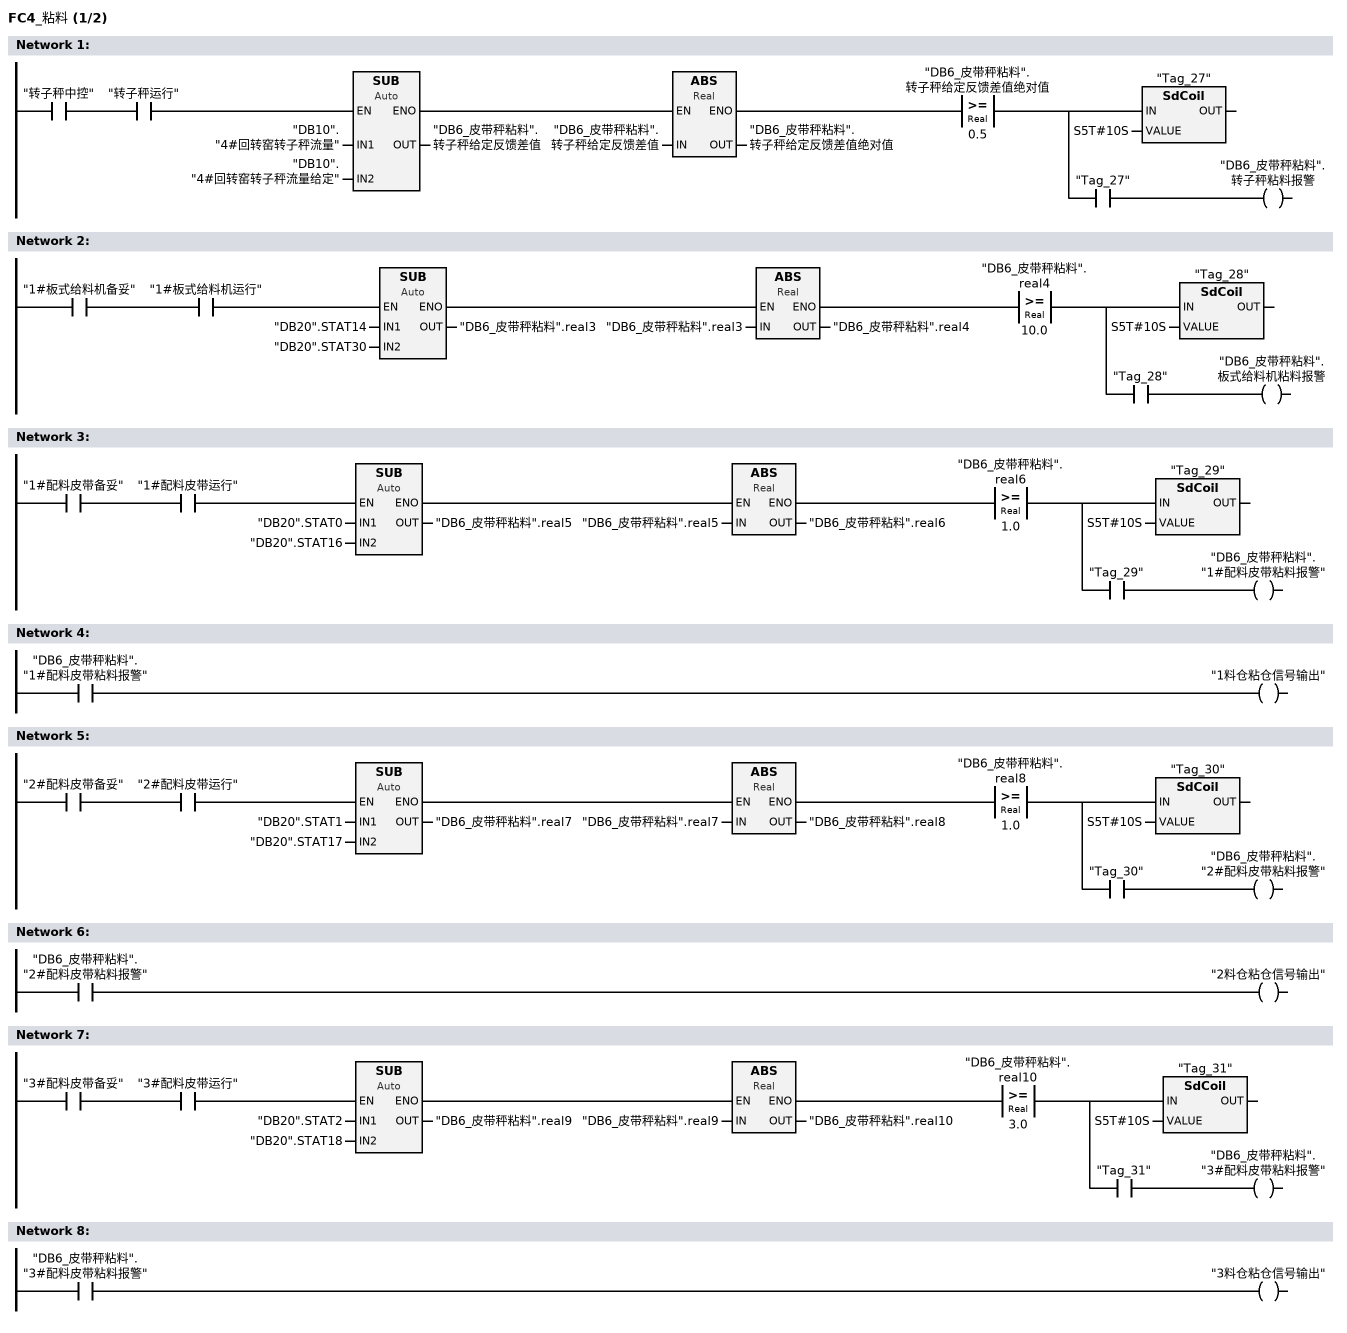
   // no SCL statement known for SdCoil: written as a call
   #_w1 := "转子秤中控" AND "转子秤运行";
   IF #_w1 THEN
       "DB6_皮带秤粘料".转子秤给定反馈差值 := "DB10"."4#回转窑转子秤流量" - "DB10"."4#回转窑转子秤流量给定";
       "DB6_皮带秤粘料".转子秤给定反馈差值绝对值 := ABS("DB6_皮带秤粘料".转子秤给定反馈差值);
   END_IF;
   #_w2 := #_w1 AND ("DB6_皮带秤粘料".转子秤给定反馈差值绝对值 >= 0.5);
   SdCoil(in := #_w2, value := S5T#10S, operand := "Tag_27");
   "DB6_皮带秤粘料".转子秤粘料报警 := #_w2 AND "Tag_27";
END_REGION

REGION Network 2
   // no SCL statement known for SdCoil: written as a call
   #_w1 := "1#板式给料机备妥" AND "1#板式给料机运行";
   IF #_w1 THEN
       "DB6_皮带秤粘料".real3 := "DB20".STAT14 - "DB20".STAT30;
       "DB6_皮带秤粘料".real4 := ABS("DB6_皮带秤粘料".real3);
   END_IF;
   #_w2 := #_w1 AND ("DB6_皮带秤粘料".real4 >= 10.0);
   SdCoil(in := #_w2, value := S5T#10S, operand := "Tag_28");
   "DB6_皮带秤粘料".板式给料机粘料报警 := #_w2 AND "Tag_28";
END_REGION

REGION Network 3
   // no SCL statement known for SdCoil: written as a call
   #_w1 := "1#配料皮带备妥" AND "1#配料皮带运行";
   IF #_w1 THEN
       "DB6_皮带秤粘料".real5 := "DB20".STAT0 - "DB20".STAT16;
       "DB6_皮带秤粘料".real6 := ABS("DB6_皮带秤粘料".real5);
   END_IF;
   #_w2 := #_w1 AND ("DB6_皮带秤粘料".real6 >= 1.0);
   SdCoil(in := #_w2, value := S5T#10S, operand := "Tag_29");
   "DB6_皮带秤粘料"."1#配料皮带粘料报警" := #_w2 AND "Tag_29";
END_REGION

REGION Network 4
   RUNG wire#powerrail
      Contact( "DB6_皮带秤粘料"."1#配料皮带粘料报警" )
      Coil( "1料仓粘仓信号输出" )
   END_RUNG
   // the same network as SCL:
   "1料仓粘仓信号输出" := "DB6_皮带秤粘料"."1#配料皮带粘料报警";
END_REGION

REGION Network 5
   // no SCL statement known for SdCoil: written as a call
   #_w1 := "2#配料皮带备妥" AND "2#配料皮带运行";
   IF #_w1 THEN
       "DB6_皮带秤粘料".real7 := "DB20".STAT1 - "DB20".STAT17;
       "DB6_皮带秤粘料".real8 := ABS("DB6_皮带秤粘料".real7);
   END_IF;
   #_w2 := #_w1 AND ("DB6_皮带秤粘料".real8 >= 1.0);
   SdCoil(in := #_w2, value := S5T#10S, operand := "Tag_30");
   "DB6_皮带秤粘料"."2#配料皮带粘料报警" := #_w2 AND "Tag_30";
END_REGION

REGION Network 6
   RUNG wire#powerrail
      Contact( "DB6_皮带秤粘料"."2#配料皮带粘料报警" )
      Coil( "2料仓粘仓信号输出" )
   END_RUNG
   // the same network as SCL:
   "2料仓粘仓信号输出" := "DB6_皮带秤粘料"."2#配料皮带粘料报警";
END_REGION

REGION Network 7
   // no SCL statement known for SdCoil: written as a call
   #_w1 := "3#配料皮带备妥" AND "3#配料皮带运行";
   IF #_w1 THEN
       "DB6_皮带秤粘料".real9 := "DB20".STAT2 - "DB20".STAT18;
       "DB6_皮带秤粘料".real10 := ABS("DB6_皮带秤粘料".real9);
   END_IF;
   #_w2 := #_w1 AND ("DB6_皮带秤粘料".real10 >= 3.0);
   SdCoil(in := #_w2, value := S5T#10S, operand := "Tag_31");
   "DB6_皮带秤粘料"."3#配料皮带粘料报警" := #_w2 AND "Tag_31";
END_REGION

REGION Network 8
   RUNG wire#powerrail
      Contact( "DB6_皮带秤粘料"."3#配料皮带粘料报警" )
      Coil( "3料仓粘仓信号输出" )
   END_RUNG
   // the same network as SCL:
   "3料仓粘仓信号输出" := "DB6_皮带秤粘料"."3#配料皮带粘料报警";
END_REGION

REGION Network 9
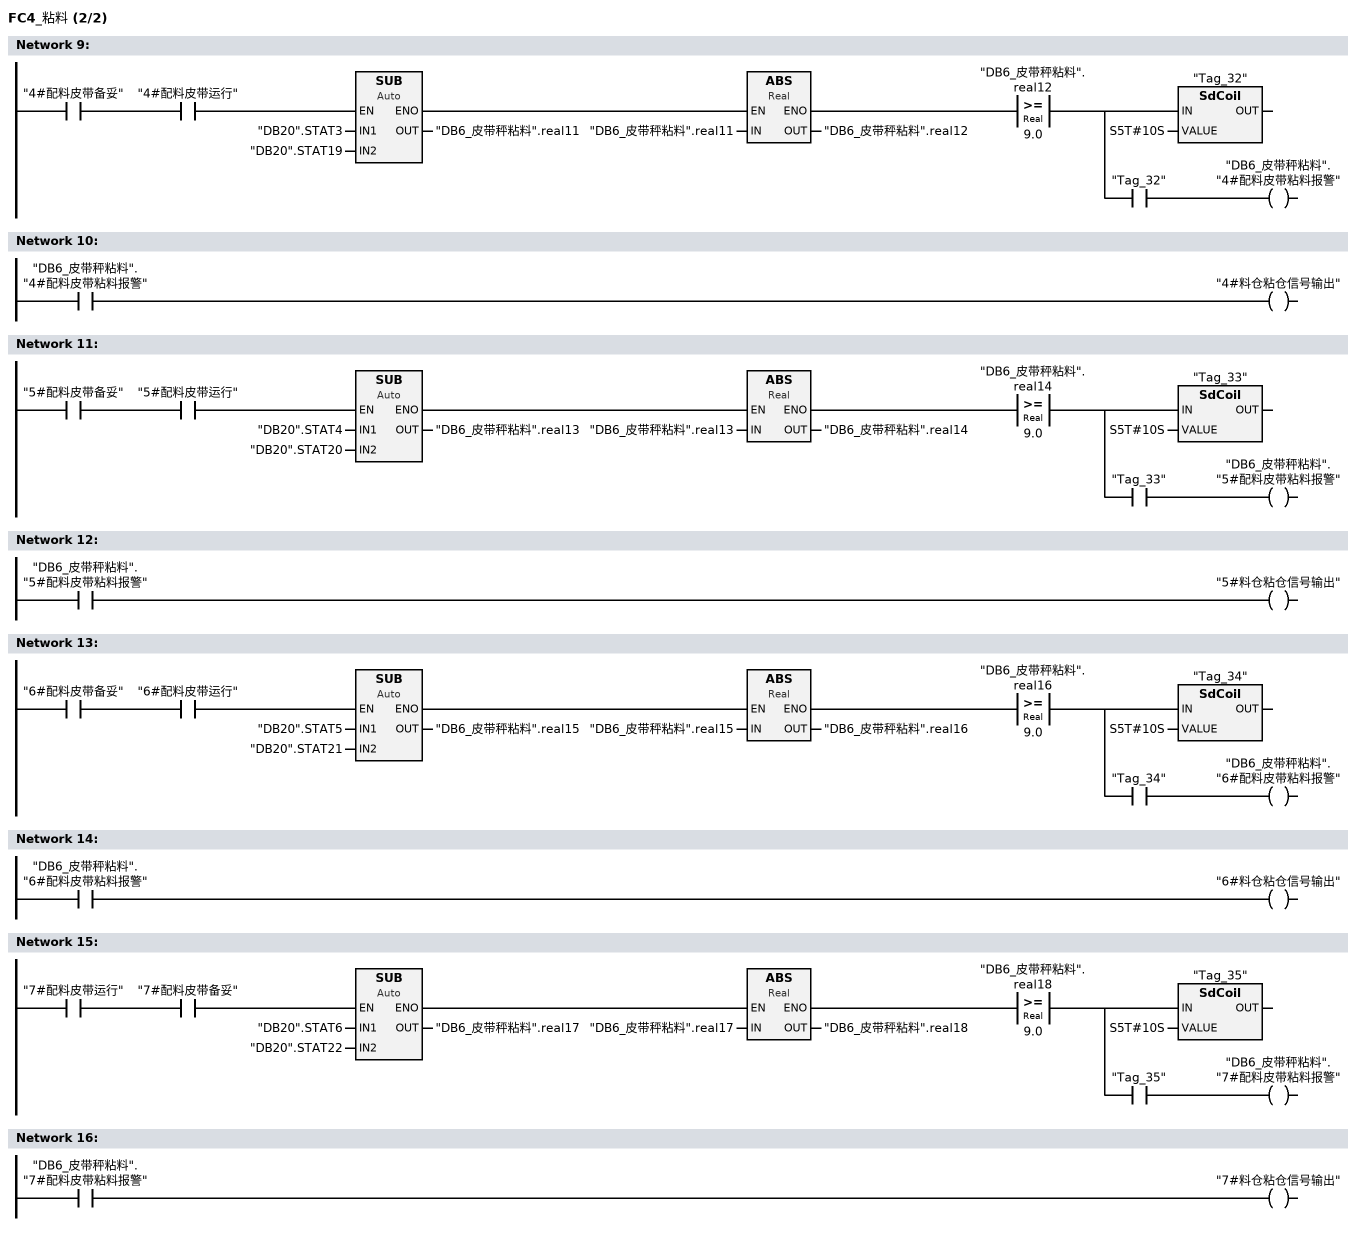
   // no SCL statement known for SdCoil: written as a call
   #_w1 := "4#配料皮带备妥" AND "4#配料皮带运行";
   IF #_w1 THEN
       "DB6_皮带秤粘料".real11 := "DB20".STAT3 - "DB20".STAT19;
       "DB6_皮带秤粘料".real12 := ABS("DB6_皮带秤粘料".real11);
   END_IF;
   #_w2 := #_w1 AND ("DB6_皮带秤粘料".real12 >= 9.0);
   SdCoil(in := #_w2, value := S5T#10S, operand := "Tag_32");
   "DB6_皮带秤粘料"."4#配料皮带粘料报警" := #_w2 AND "Tag_32";
END_REGION

REGION Network 10
   RUNG wire#powerrail
      Contact( "DB6_皮带秤粘料"."4#配料皮带粘料报警" )
      Coil( "4#料仓粘仓信号输出" )
   END_RUNG
   // the same network as SCL:
   "4#料仓粘仓信号输出" := "DB6_皮带秤粘料"."4#配料皮带粘料报警";
END_REGION

REGION Network 11
   // no SCL statement known for SdCoil: written as a call
   #_w1 := "5#配料皮带备妥" AND "5#配料皮带运行";
   IF #_w1 THEN
       "DB6_皮带秤粘料".real13 := "DB20".STAT4 - "DB20".STAT20;
       "DB6_皮带秤粘料".real14 := ABS("DB6_皮带秤粘料".real13);
   END_IF;
   #_w2 := #_w1 AND ("DB6_皮带秤粘料".real14 >= 9.0);
   SdCoil(in := #_w2, value := S5T#10S, operand := "Tag_33");
   "DB6_皮带秤粘料"."5#配料皮带粘料报警" := #_w2 AND "Tag_33";
END_REGION

REGION Network 12
   RUNG wire#powerrail
      Contact( "DB6_皮带秤粘料"."5#配料皮带粘料报警" )
      Coil( "5#料仓粘仓信号输出" )
   END_RUNG
   // the same network as SCL:
   "5#料仓粘仓信号输出" := "DB6_皮带秤粘料"."5#配料皮带粘料报警";
END_REGION

REGION Network 13
   // no SCL statement known for SdCoil: written as a call
   #_w1 := "6#配料皮带备妥" AND "6#配料皮带运行";
   IF #_w1 THEN
       "DB6_皮带秤粘料".real15 := "DB20".STAT5 - "DB20".STAT21;
       "DB6_皮带秤粘料".real16 := ABS("DB6_皮带秤粘料".real15);
   END_IF;
   #_w2 := #_w1 AND ("DB6_皮带秤粘料".real16 >= 9.0);
   SdCoil(in := #_w2, value := S5T#10S, operand := "Tag_34");
   "DB6_皮带秤粘料"."6#配料皮带粘料报警" := #_w2 AND "Tag_34";
END_REGION

REGION Network 14
   RUNG wire#powerrail
      Contact( "DB6_皮带秤粘料"."6#配料皮带粘料报警" )
      Coil( "6#料仓粘仓信号输出" )
   END_RUNG
   // the same network as SCL:
   "6#料仓粘仓信号输出" := "DB6_皮带秤粘料"."6#配料皮带粘料报警";
END_REGION

REGION Network 15
   // no SCL statement known for SdCoil: written as a call
   #_w1 := "7#配料皮带运行" AND "7#配料皮带备妥";
   IF #_w1 THEN
       "DB6_皮带秤粘料".real17 := "DB20".STAT6 - "DB20".STAT22;
       "DB6_皮带秤粘料".real18 := ABS("DB6_皮带秤粘料".real17);
   END_IF;
   #_w2 := #_w1 AND ("DB6_皮带秤粘料".real18 >= 9.0);
   SdCoil(in := #_w2, value := S5T#10S, operand := "Tag_35");
   "DB6_皮带秤粘料"."7#配料皮带粘料报警" := #_w2 AND "Tag_35";
END_REGION

REGION Network 16
   RUNG wire#powerrail
      Contact( "DB6_皮带秤粘料"."7#配料皮带粘料报警" )
      Coil( "7#料仓粘仓信号输出" )
   END_RUNG
   // the same network as SCL:
   "7#料仓粘仓信号输出" := "DB6_皮带秤粘料"."7#配料皮带粘料报警";
END_REGION
END_FUNCTION

FUNCTION "回转窑控制" : Void   // FC11, LAD
{ S7_Optimized_Access := 'FALSE' }
VERSION : 0.1
   VAR_TEMP   // added for the SCL form of the ladder/FBD networks
      _w1 : Bool;
      _s5time1 : S5Time;
   END_VAR
BEGIN

REGION Network 1
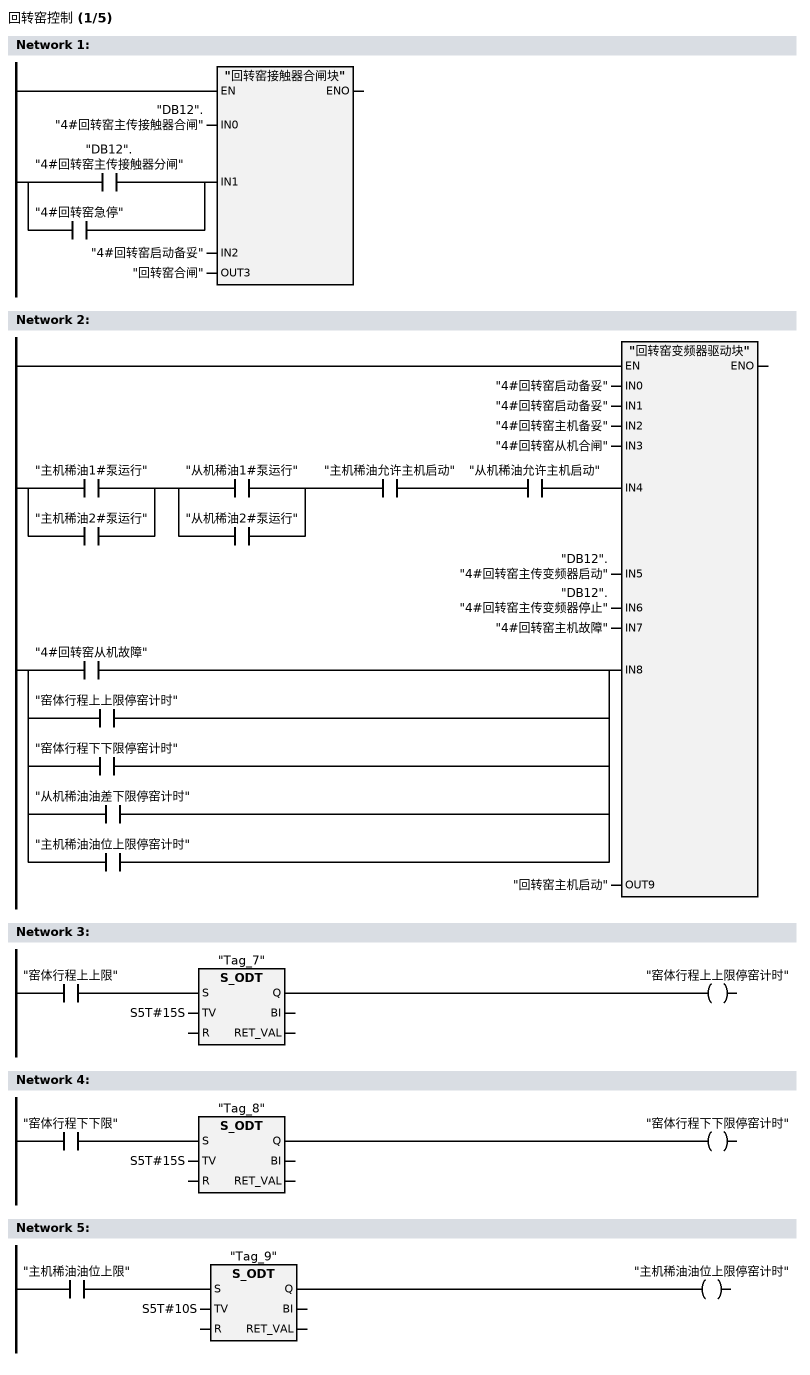
   RUNG wire#powerrail
      "回转窑接触器合闸块"(IN1 := wire#w1, IN0 := "DB12"."4#回转窑主传接触器合闸", IN2 := "4#回转窑启动备妥", OUT3 := "回转窑合闸")
   END_RUNG
   RUNG wire#powerrail
      Contact( "DB12"."4#回转窑主传接触器分闸" )
   END_RUNG wire#w1
   RUNG wire#powerrail
      Contact( "4#回转窑急停" )
   END_RUNG wire#w1
   // the same network as SCL:
   "回转窑接触器合闸块"(IN0 := "DB12"."4#回转窑主传接触器合闸",
               IN1 := "DB12"."4#回转窑主传接触器分闸" OR "4#回转窑急停",
               IN2 := "4#回转窑启动备妥",
               OUT3 := "回转窑合闸");
END_REGION

REGION Network 2
   RUNG wire#powerrail
      "回转窑变频器驱动块"(IN4 := wire#w3, IN8 := wire#w4, IN0 := "4#回转窑启动备妥", IN1 := "4#回转窑启动备妥", IN2 := "4#回转窑主机备妥", IN3 := "4#回转窑从机合闸", IN5 := "DB12"."4#回转窑主传变频器启动", IN6 := "DB12"."4#回转窑主传变频器停止", IN7 := "4#回转窑主机故障", OUT9 := "回转窑主机启动")
   END_RUNG
   RUNG wire#powerrail
      Contact( "主机稀油1#泵运行" )
      wire#w1
      Contact( "从机稀油1#泵运行" )
      wire#w2
      Contact( "主机稀油允许主机启动" )
      Contact( "从机稀油允许主机启动" )
   END_RUNG wire#w3
   RUNG wire#powerrail
      Contact( "主机稀油2#泵运行" )
   END_RUNG wire#w1
   RUNG wire#w1
      Contact( "从机稀油2#泵运行" )
   END_RUNG wire#w2
   RUNG wire#powerrail
      Contact( "4#回转窑从机故障" )
   END_RUNG wire#w4
   RUNG wire#powerrail
      Contact( "窑体行程上上限停窑计时" )
   END_RUNG wire#w4
   RUNG wire#powerrail
      Contact( "窑体行程下下限停窑计时" )
   END_RUNG wire#w4
   RUNG wire#powerrail
      Contact( "从机稀油油差下限停窑计时" )
   END_RUNG wire#w4
   RUNG wire#powerrail
      Contact( "主机稀油油位上限停窑计时" )
   END_RUNG wire#w4
   // the same network as SCL:
   "回转窑变频器驱动块"(IN0 := "4#回转窑启动备妥",
               IN1 := "4#回转窑启动备妥",
               IN2 := "4#回转窑主机备妥",
               IN3 := "4#回转窑从机合闸",
               IN4 := ("主机稀油1#泵运行" OR "主机稀油2#泵运行") AND ("从机稀油1#泵运行" OR "从机稀油2#泵运行") AND "主机稀油允许主机启动" AND "从机稀油允许主机启动",
               IN5 := "DB12"."4#回转窑主传变频器启动",
               IN6 := "DB12"."4#回转窑主传变频器停止",
               IN7 := "4#回转窑主机故障",
               IN8 := "4#回转窑从机故障" OR "窑体行程上上限停窑计时" OR "窑体行程下下限停窑计时" OR "从机稀油油差下限停窑计时" OR "主机稀油油位上限停窑计时",
               OUT9 := "回转窑主机启动");
END_REGION

REGION Network 3
   RUNG wire#powerrail
      Contact( "窑体行程上上限" )
      S_ODT(T_NO := "Tag_7", TV := S5T#15S, R :=, BI =>, RET_VAL =>)
      Coil( "窑体行程上上限停窑计时" )
   END_RUNG
   // the same network as SCL:
   #_s5time1 := S_ODT(T_NO := "Tag_7", TV := S5T#15S, S := "窑体行程上上限", Q => #_w1);
   "窑体行程上上限停窑计时" := #_w1;
END_REGION

REGION Network 4
   RUNG wire#powerrail
      Contact( "窑体行程下下限" )
      S_ODT(T_NO := "Tag_8", TV := S5T#15S, R :=, BI =>, RET_VAL =>)
      Coil( "窑体行程下下限停窑计时" )
   END_RUNG
   // the same network as SCL:
   #_s5time1 := S_ODT(T_NO := "Tag_8", TV := S5T#15S, S := "窑体行程下下限", Q => #_w1);
   "窑体行程下下限停窑计时" := #_w1;
END_REGION

REGION Network 5
   RUNG wire#powerrail
      Contact( "主机稀油油位上限" )
      S_ODT(T_NO := "Tag_9", TV := S5T#10S, R :=, BI =>, RET_VAL =>)
      Coil( "主机稀油油位上限停窑计时" )
   END_RUNG
   // the same network as SCL:
   #_s5time1 := S_ODT(T_NO := "Tag_9", S := "主机稀油油位上限", TV := S5T#10S, Q => #_w1);
   "主机稀油油位上限停窑计时" := #_w1;
END_REGION

REGION Network 6
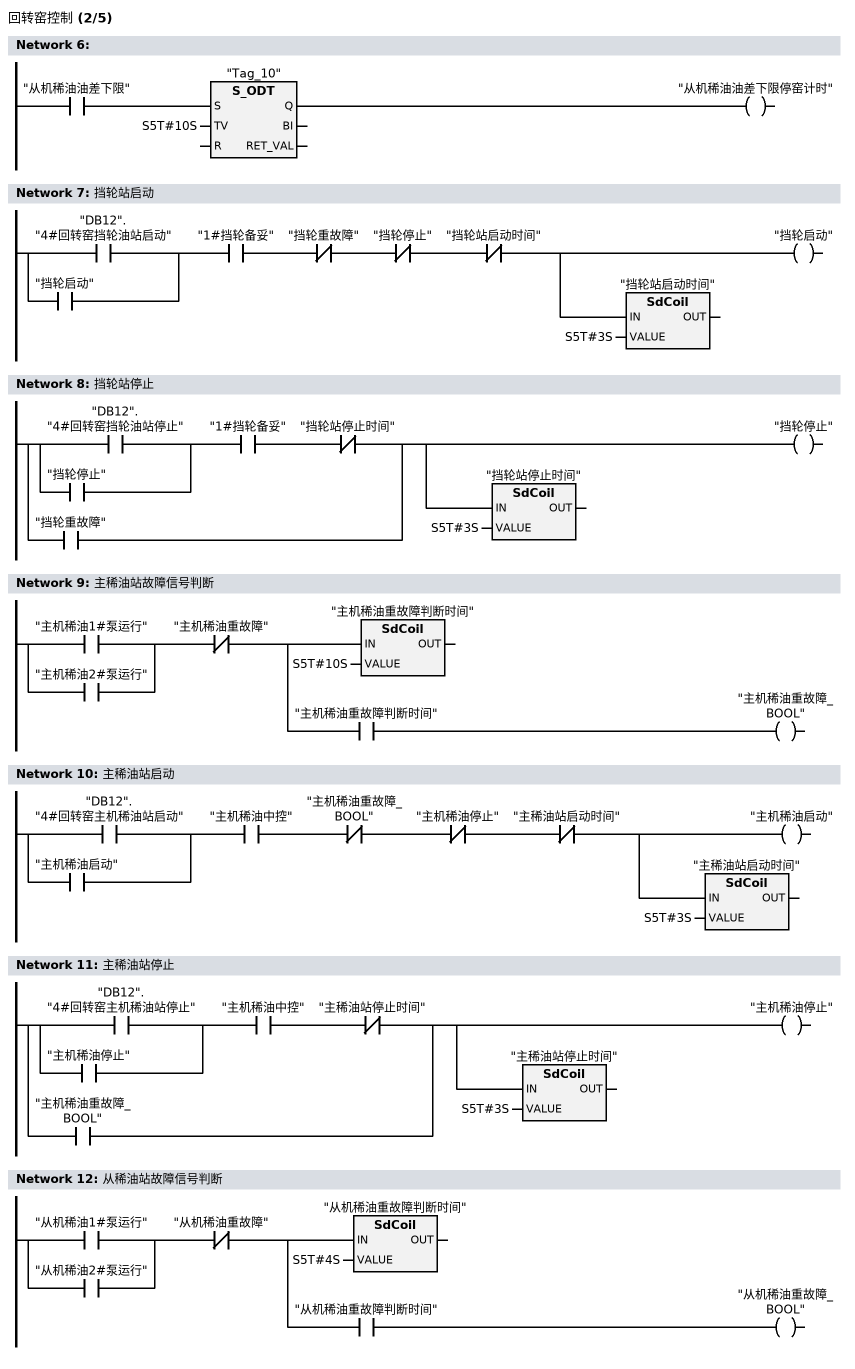
   RUNG wire#powerrail
      Contact( "从机稀油油差下限" )
      S_ODT(T_NO := "Tag_10", TV := S5T#10S, R :=, BI =>, RET_VAL =>)
      Coil( "从机稀油油差下限停窑计时" )
   END_RUNG
   // the same network as SCL:
   #_s5time1 := S_ODT(T_NO := "Tag_10", TV := S5T#10S, S := "从机稀油油差下限", Q => #_w1);
   "从机稀油油差下限停窑计时" := #_w1;
END_REGION

REGION Network 7: 挡轮站启动
   // no SCL statement known for SdCoil: written as a call
   "挡轮启动" := ("DB12"."4#回转窑挡轮油站启动" OR "挡轮启动") AND "1#挡轮备妥" AND NOT "挡轮重故障" AND NOT "挡轮停止" AND NOT "挡轮站启动时间";
   SdCoil(in := "挡轮启动", value := S5T#3S, operand := "挡轮站启动时间");
END_REGION

REGION Network 8: 挡轮站停止
   // no SCL statement known for SdCoil: written as a call
   "挡轮停止" := (("DB12"."4#回转窑挡轮油站停止" OR "挡轮停止") AND "1#挡轮备妥" AND NOT "挡轮站停止时间") OR "挡轮重故障";
   SdCoil(in := "挡轮停止", value := S5T#3S, operand := "挡轮站停止时间");
END_REGION

REGION Network 9: 主稀油站故障信号判断
   // no SCL statement known for SdCoil: written as a call
   #_w1 := ("主机稀油1#泵运行" OR "主机稀油2#泵运行") AND NOT "主机稀油重故障";
   SdCoil(in := #_w1, value := S5T#10S, operand := "主机稀油重故障判断时间");
   "主机稀油重故障_BOOL" := #_w1 AND "主机稀油重故障判断时间";
END_REGION

REGION Network 10: 主稀油站启动
   // no SCL statement known for SdCoil: written as a call
   "主机稀油启动" := ("DB12"."4#回转窑主机稀油站启动" OR "主机稀油启动") AND "主机稀油中控" AND NOT "主机稀油重故障_BOOL" AND NOT "主机稀油停止" AND NOT "主稀油站启动时间";
   SdCoil(in := "主机稀油启动", value := S5T#3S, operand := "主稀油站启动时间");
END_REGION

REGION Network 11: 主稀油站停止
   // no SCL statement known for SdCoil: written as a call
   "主机稀油停止" := (("DB12"."4#回转窑主机稀油站停止" OR "主机稀油停止") AND "主机稀油中控" AND NOT "主稀油站停止时间") OR "主机稀油重故障_BOOL";
   SdCoil(in := "主机稀油停止", value := S5T#3S, operand := "主稀油站停止时间");
END_REGION

REGION Network 12: 从稀油站故障信号判断
   // no SCL statement known for SdCoil: written as a call
   #_w1 := ("从机稀油1#泵运行" OR "从机稀油2#泵运行") AND NOT "从机稀油重故障";
   SdCoil(in := #_w1, value := S5T#4S, operand := "从机稀油重故障判断时间");
   "从机稀油重故障_BOOL" := #_w1 AND "从机稀油重故障判断时间";
END_REGION

REGION Network 13: 从稀油站启动
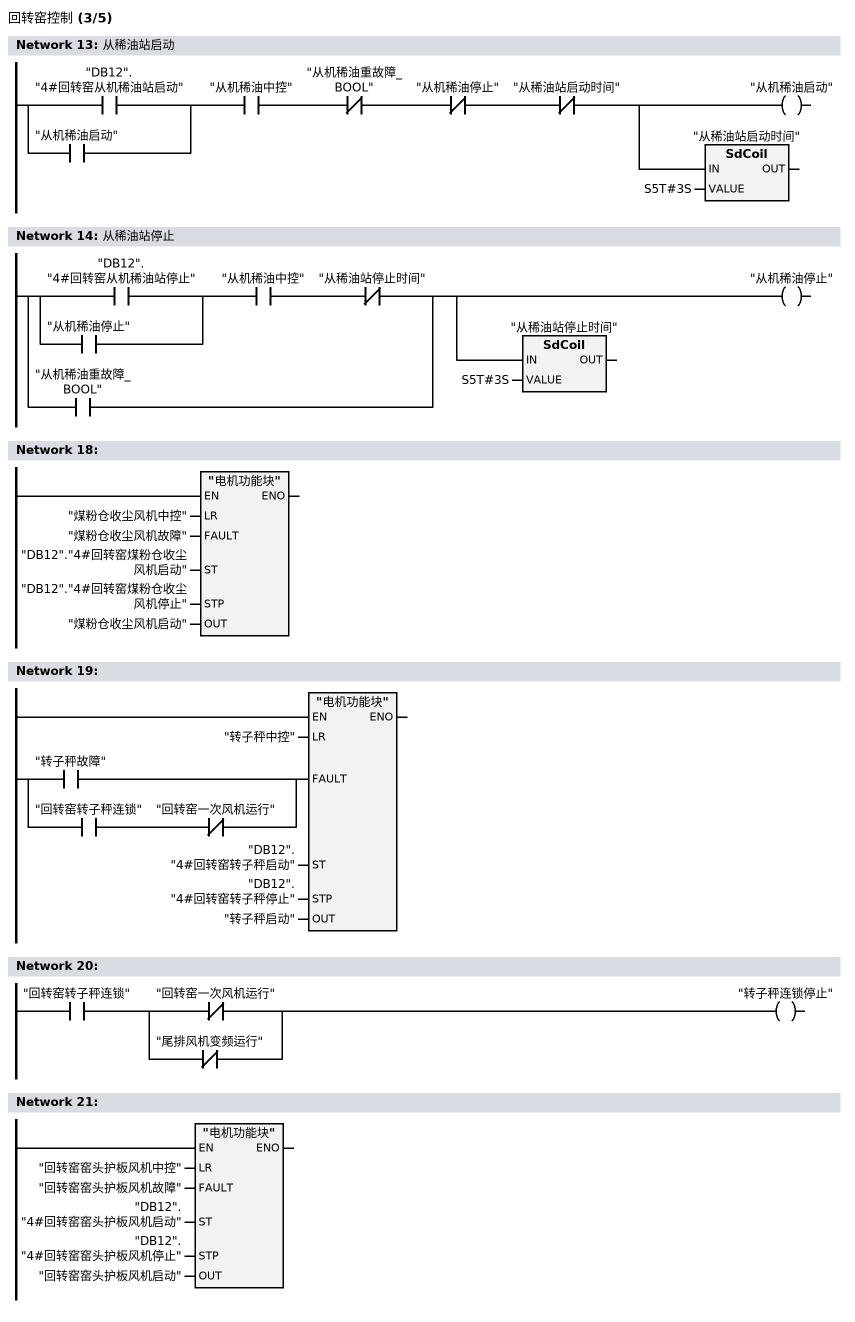
   // no SCL statement known for SdCoil: written as a call
   "从机稀油启动" := ("DB12"."4#回转窑从机稀油站启动" OR "从机稀油启动") AND "从机稀油中控" AND NOT "从机稀油重故障_BOOL" AND NOT "从机稀油停止" AND NOT "从稀油站启动时间";
   SdCoil(in := "从机稀油启动", value := S5T#3S, operand := "从稀油站启动时间");
END_REGION

REGION Network 14: 从稀油站停止
   // no SCL statement known for SdCoil: written as a call
   "从机稀油停止" := (("DB12"."4#回转窑从机稀油站停止" OR "从机稀油停止") AND "从机稀油中控" AND NOT "从稀油站停止时间") OR "从机稀油重故障_BOOL";
   SdCoil(in := "从机稀油停止", value := S5T#3S, operand := "从稀油站停止时间");
END_REGION

REGION Network 18
   RUNG wire#powerrail
      "电机功能块"(LR := "煤粉仓收尘风机中控", FAULT := "煤粉仓收尘风机故障", ST := "DB12"."4#回转窑煤粉仓收尘风机启动", STP := "DB12"."4#回转窑煤粉仓收尘风机停止", OUT := "煤粉仓收尘风机启动")
   END_RUNG
   // the same network as SCL:
   "电机功能块"(LR := "煤粉仓收尘风机中控",
           FAULT := "煤粉仓收尘风机故障",
           ST := "DB12"."4#回转窑煤粉仓收尘风机启动",
           STP := "DB12"."4#回转窑煤粉仓收尘风机停止",
           OUT := "煤粉仓收尘风机启动");
END_REGION

REGION Network 19
   RUNG wire#powerrail
      "电机功能块"(FAULT := wire#w1, LR := "转子秤中控", ST := "DB12"."4#回转窑转子秤启动", STP := "DB12"."4#回转窑转子秤停止", OUT := "转子秤启动")
   END_RUNG
   RUNG wire#powerrail
      Contact( "转子秤故障" )
   END_RUNG wire#w1
   RUNG wire#powerrail
      Contact( "回转窑转子秤连锁" )
      I_Contact( "回转窑一次风机运行" )
   END_RUNG wire#w1
   // the same network as SCL:
   "电机功能块"(LR := "转子秤中控",
           FAULT := "转子秤故障" OR ("回转窑转子秤连锁" AND NOT "回转窑一次风机运行"),
           ST := "DB12"."4#回转窑转子秤启动",
           STP := "DB12"."4#回转窑转子秤停止",
           OUT := "转子秤启动");
END_REGION

REGION Network 20
   RUNG wire#powerrail
      Contact( "回转窑转子秤连锁" )
      wire#w1
      I_Contact( "回转窑一次风机运行" )
      wire#w2
      Coil( "转子秤连锁停止" )
   END_RUNG
   RUNG wire#w1
      I_Contact( "尾排风机变频运行" )
   END_RUNG wire#w2
   // the same network as SCL:
   "转子秤连锁停止" := "回转窑转子秤连锁" AND (NOT "回转窑一次风机运行" OR NOT "尾排风机变频运行");
END_REGION

REGION Network 21
   RUNG wire#powerrail
      "电机功能块"(LR := "回转窑窑头护板风机中控", FAULT := "回转窑窑头护板风机故障", ST := "DB12"."4#回转窑窑头护板风机启动", STP := "DB12"."4#回转窑窑头护板风机停止", OUT := "回转窑窑头护板风机启动")
   END_RUNG
   // the same network as SCL:
   "电机功能块"(LR := "回转窑窑头护板风机中控",
           FAULT := "回转窑窑头护板风机故障",
           ST := "DB12"."4#回转窑窑头护板风机启动",
           STP := "DB12"."4#回转窑窑头护板风机停止",
           OUT := "回转窑窑头护板风机启动");
END_REGION

REGION Network 22
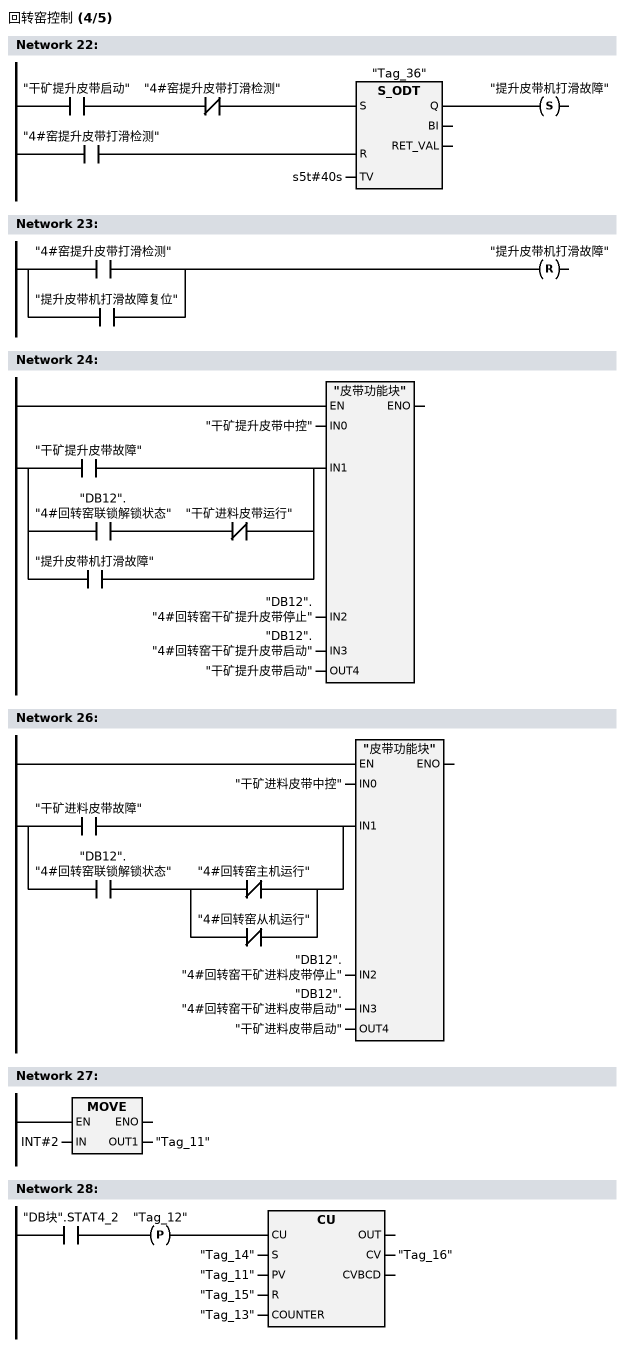
   RUNG wire#powerrail
      Contact( "干矿提升皮带启动" )
      I_Contact( "4#窑提升皮带打滑检测" )
      S_ODT(T_NO := "Tag_36", R := wire#w1, TV := s5t#40s, BI =>, RET_VAL =>)
      S_Coil( "提升皮带机打滑故障" )
   END_RUNG
   RUNG wire#powerrail
      Contact( "4#窑提升皮带打滑检测" )
   END_RUNG wire#w1
   // the same network as SCL:
   #_s5time1 := S_ODT(T_NO := "Tag_36",
                      S := "干矿提升皮带启动" AND NOT "4#窑提升皮带打滑检测",
                      R := "4#窑提升皮带打滑检测",
                      TV := s5t#40s,
                      Q => #_w1);
   IF #_w1 THEN "提升皮带机打滑故障" := TRUE; END_IF;
END_REGION

REGION Network 23
   RUNG wire#powerrail
      Contact( "4#窑提升皮带打滑检测" )
      wire#w1
      R_Coil( "提升皮带机打滑故障" )
   END_RUNG
   RUNG wire#powerrail
      Contact( "提升皮带机打滑故障复位" )
   END_RUNG wire#w1
   // the same network as SCL:
   IF "4#窑提升皮带打滑检测" OR "提升皮带机打滑故障复位" THEN "提升皮带机打滑故障" := FALSE; END_IF;
END_REGION

REGION Network 24
   RUNG wire#powerrail
      "皮带功能块"(IN1 := wire#w1, IN0 := "干矿提升皮带中控", IN2 := "DB12"."4#回转窑干矿提升皮带停止", IN3 := "DB12"."4#回转窑干矿提升皮带启动", OUT4 := "干矿提升皮带启动")
   END_RUNG
   RUNG wire#powerrail
      Contact( "干矿提升皮带故障" )
   END_RUNG wire#w1
   RUNG wire#powerrail
      Contact( "DB12"."4#回转窑联锁解锁状态" )
      I_Contact( "干矿进料皮带运行" )
   END_RUNG wire#w1
   RUNG wire#powerrail
      Contact( "提升皮带机打滑故障" )
   END_RUNG wire#w1
   // the same network as SCL:
   "皮带功能块"(IN0 := "干矿提升皮带中控",
           IN1 := "干矿提升皮带故障" OR ("DB12"."4#回转窑联锁解锁状态" AND NOT "干矿进料皮带运行") OR "提升皮带机打滑故障",
           IN2 := "DB12"."4#回转窑干矿提升皮带停止",
           IN3 := "DB12"."4#回转窑干矿提升皮带启动",
           OUT4 := "干矿提升皮带启动");
END_REGION

REGION Network 26
   RUNG wire#powerrail
      "皮带功能块"(IN1 := wire#w2, IN0 := "干矿进料皮带中控", IN2 := "DB12"."4#回转窑干矿进料皮带停止", IN3 := "DB12"."4#回转窑干矿进料皮带启动", OUT4 := "干矿进料皮带启动")
   END_RUNG
   RUNG wire#powerrail
      Contact( "干矿进料皮带故障" )
   END_RUNG wire#w2
   RUNG wire#powerrail
      Contact( "DB12"."4#回转窑联锁解锁状态" )
      wire#w1
      I_Contact( "4#回转窑主机运行" )
   END_RUNG wire#w2
   RUNG wire#w1
      I_Contact( "4#回转窑从机运行" )
   END_RUNG wire#w2
   // the same network as SCL:
   "皮带功能块"(IN0 := "干矿进料皮带中控",
           IN1 := "干矿进料皮带故障" OR ("DB12"."4#回转窑联锁解锁状态" AND (NOT "4#回转窑主机运行" OR NOT "4#回转窑从机运行")),
           IN2 := "DB12"."4#回转窑干矿进料皮带停止",
           IN3 := "DB12"."4#回转窑干矿进料皮带启动",
           OUT4 := "干矿进料皮带启动");
END_REGION

REGION Network 27
   RUNG wire#powerrail
      { S7_GenerateENO := "TRUE" } Move(in := INT#2, out1 => "Tag_11")
   END_RUNG
   // the same network as SCL:
   "Tag_11" := INT#2;
END_REGION

REGION Network 28
   // no SCL statement known for Cu: written as a call
   #_w1 := "DB块".STAT4_2 AND NOT "Tag_12";   // rising edge
   "Tag_12" := "DB块".STAT4_2;
   Cu(cu := #_w1, s := "Tag_14", pv := "Tag_11", r := "Tag_15", "counter" := "Tag_13", cv => "Tag_16");
END_REGION

REGION Network 29
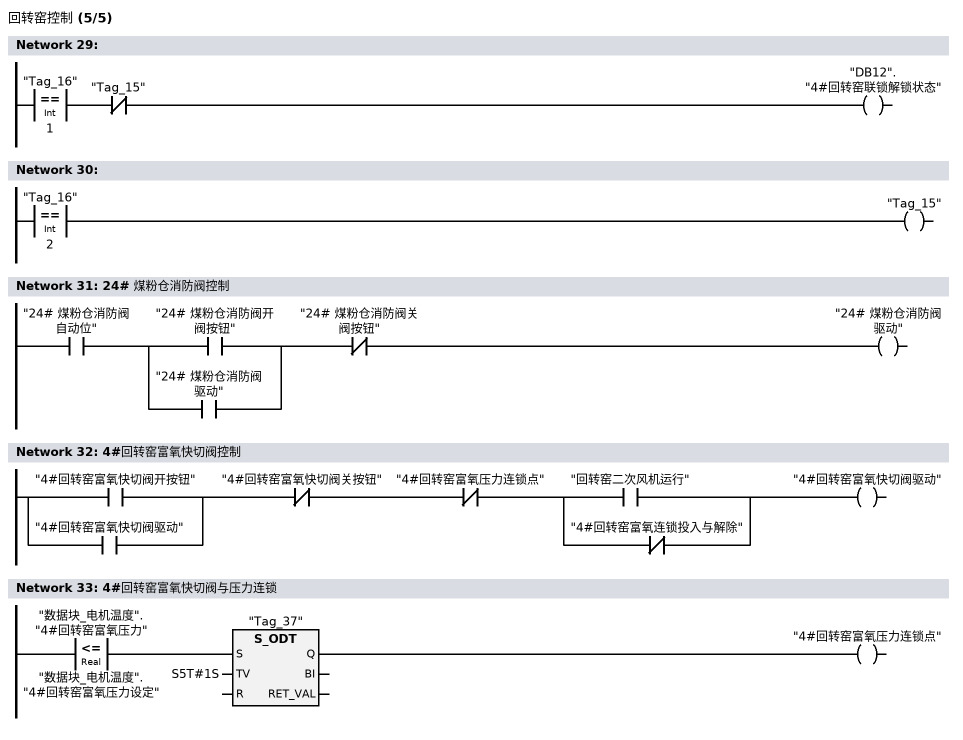
   RUNG wire#powerrail
      { S7_Templates := "SrcType := Int" } EQ_Contact(in1 := "Tag_16", in2 := 1)
      I_Contact( "Tag_15" )
      Coil( "DB12"."4#回转窑联锁解锁状态" )
   END_RUNG
   // the same network as SCL:
   "DB12"."4#回转窑联锁解锁状态" := ("Tag_16" = 1) AND NOT "Tag_15";
END_REGION

REGION Network 30
   RUNG wire#powerrail
      { S7_Templates := "SrcType := Int" } EQ_Contact(in1 := "Tag_16", in2 := 2)
      Coil( "Tag_15" )
   END_RUNG
   // the same network as SCL:
   "Tag_15" := "Tag_16" = 2;
END_REGION

REGION Network 31: 24# 煤粉仓消防阀控制
   RUNG wire#powerrail
      Contact( "24# 煤粉仓消防阀自动位" )
      wire#w1
      Contact( "24# 煤粉仓消防阀开阀按钮" )
      wire#w2
      I_Contact( "24# 煤粉仓消防阀关阀按钮" )
      Coil( "24# 煤粉仓消防阀驱动" )
   END_RUNG
   RUNG wire#w1
      Contact( "24# 煤粉仓消防阀驱动" )
   END_RUNG wire#w2
   // the same network as SCL:
   "24# 煤粉仓消防阀驱动" := "24# 煤粉仓消防阀自动位" AND ("24# 煤粉仓消防阀开阀按钮" OR "24# 煤粉仓消防阀驱动") AND NOT "24# 煤粉仓消防阀关阀按钮";
END_REGION

REGION Network 32: 4#回转窑富氧快切阀控制
   RUNG wire#powerrail
      Contact( "4#回转窑富氧快切阀开按钮" )
      wire#w1
      I_Contact( "4#回转窑富氧快切阀关按钮" )
      I_Contact( "4#回转窑富氧压力连锁点" )
      wire#w2
      Contact( "回转窑二次风机运行" )
      wire#w3
      Coil( "4#回转窑富氧快切阀驱动" )
   END_RUNG
   RUNG wire#powerrail
      Contact( "4#回转窑富氧快切阀驱动" )
   END_RUNG wire#w1
   RUNG wire#w2
      I_Contact( "4#回转窑富氧连锁投入与解除" )
   END_RUNG wire#w3
   // the same network as SCL:
   "4#回转窑富氧快切阀驱动" := ("4#回转窑富氧快切阀开按钮" OR "4#回转窑富氧快切阀驱动") AND NOT "4#回转窑富氧快切阀关按钮" AND NOT "4#回转窑富氧压力连锁点" AND ("回转窑二次风机运行" OR NOT "4#回转窑富氧连锁投入与解除");
END_REGION

REGION Network 33: 4#回转窑富氧快切阀与压力连锁
   RUNG wire#powerrail
      { S7_Templates := "SrcType := Real" } LE_Contact(in1 := "数据块_电机温度"."4#回转窑富氧压力", in2 := "数据块_电机温度"."4#回转窑富氧压力设定")
      S_ODT(T_NO := "Tag_37", TV := S5T#1S, R :=, BI =>, RET_VAL =>)
      Coil( "4#回转窑富氧压力连锁点" )
   END_RUNG
   // the same network as SCL:
   #_s5time1 := S_ODT(T_NO := "Tag_37",
                      S := "数据块_电机温度"."4#回转窑富氧压力" <= "数据块_电机温度"."4#回转窑富氧压力设定",
                      TV := S5T#1S,
                      Q => #_w1);
   "4#回转窑富氧压力连锁点" := #_w1;
END_REGION
END_FUNCTION

FUNCTION "回转窑模拟量反馈" : Void   // FC12, LAD
{ S7_Optimized_Access := 'FALSE' }
VERSION : 0.1
   VAR_TEMP   // added for the SCL form of the ladder/FBD networks
      _w1 : Bool;
      _s5time1 : S5Time;
   END_VAR
BEGIN

REGION Network 1
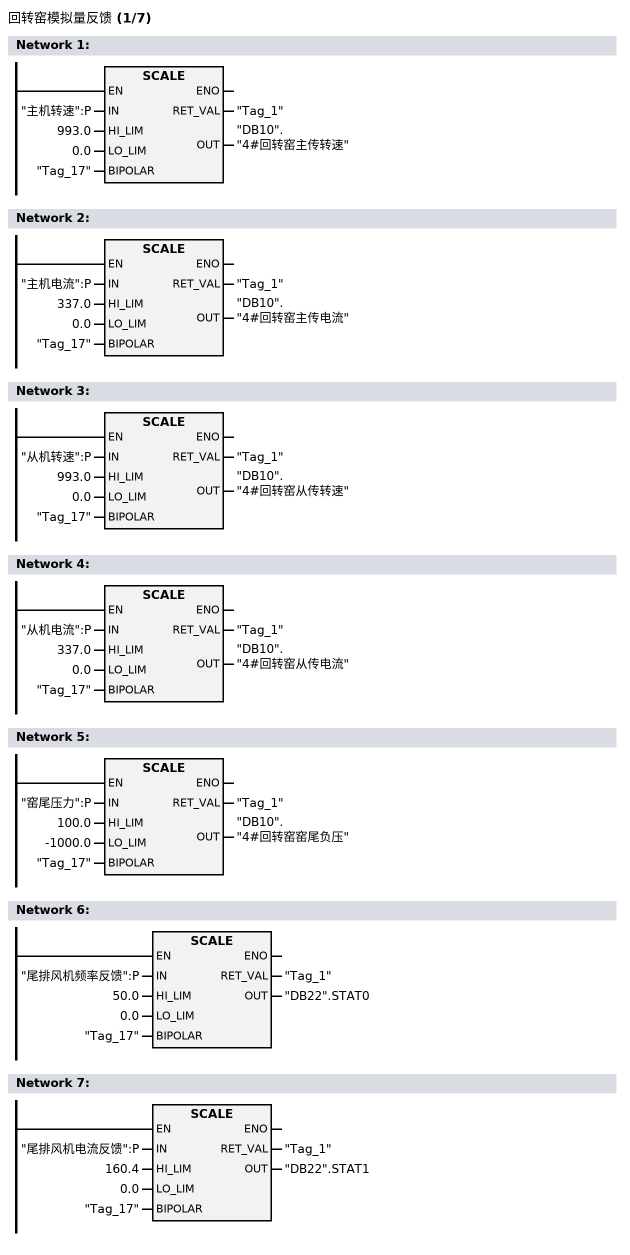
   "Tag_1" := SCALE(IN := "主机转速":P,
                    HI_LIM := 993.0,
                    LO_LIM := 0.0,
                    BIPOLAR := "Tag_17",
                    OUT => "DB10"."4#回转窑主传转速");
END_REGION

REGION Network 2
   "Tag_1" := SCALE(IN := "主机电流":P,
                    HI_LIM := 337.0,
                    LO_LIM := 0.0,
                    BIPOLAR := "Tag_17",
                    OUT => "DB10"."4#回转窑主传电流");
END_REGION

REGION Network 3
   "Tag_1" := SCALE(IN := "从机转速":P,
                    HI_LIM := 993.0,
                    LO_LIM := 0.0,
                    BIPOLAR := "Tag_17",
                    OUT => "DB10"."4#回转窑从传转速");
END_REGION

REGION Network 4
   "Tag_1" := SCALE(IN := "从机电流":P,
                    HI_LIM := 337.0,
                    LO_LIM := 0.0,
                    BIPOLAR := "Tag_17",
                    OUT => "DB10"."4#回转窑从传电流");
END_REGION

REGION Network 5
   "Tag_1" := SCALE(IN := "窑尾压力":P,
                    HI_LIM := 100.0,
                    LO_LIM := -1000.0,
                    BIPOLAR := "Tag_17",
                    OUT => "DB10"."4#回转窑窑尾负压");
END_REGION

REGION Network 6
   "Tag_1" := SCALE(IN := "尾排风机频率反馈":P, HI_LIM := 50.0, LO_LIM := 0.0, BIPOLAR := "Tag_17", OUT => "DB22".STAT0);
END_REGION

REGION Network 7
   "Tag_1" := SCALE(IN := "尾排风机电流反馈":P,
                    HI_LIM := 160.4,
                    LO_LIM := 0.0,
                    BIPOLAR := "Tag_17",
                    OUT => "DB22".STAT1);
END_REGION

REGION Network 8
